(* Logix 5000 project; controller _GigaDiscovery vendor 1 type 14 code 244 rev 35.11; software revision 35.03 *)

TASK _10_milli_sec (periodic, rate 10 ms, priority 5, watchdog 500 ms) : Main10ms
TASK MainTask (continuous, watchdog 500 ms) : Input, Alarms, General, Pylon, Recipe, Output, HMI, Restraints
TASK Pylon_Control (periodic, rate 5 ms, priority 2, watchdog 500 ms) : Pylon_Oscillation
TASK SafetyTask (periodic, rate 40 ms, priority 2, watchdog 20 ms) : S_Input, S_Alarms, S_Cycles, S_Platform_and_Gates, S_Restraints_Release, S_Output

MODULES
   Local : vendor 1 type 14 code 244 (5069 0, rev 35.11)
      Gondola_Motor_7 : vendor 1 type 152 code 121 (Ethernet 192.168.1.63, rev 7.3, Output RPI 20 ms)
           K205_MCC:12:I.4   // Compressor Motor Protection Feedback -F18002C
           K205_MCC:12:I.3   // Compressor Motor Command Feedback -F18101E
           K205_MCC:12:I.2   // Motor 7 Thermal Probe -K16602H
           K205_MCC:12:I.1   // Motor 7 Fan Protection Feedback -F16402C
           K205_MCC:12:I.0   // Zero Set Sensor -B11201A
           K205_MCC:12:I.6   // Platform closed Sector 1 -B22501J
           K205_MCC:12:I.5   // Dryer Motor Protection Feedback -F18202C
           K205_MCC:12:I.7   // Platform closed Sector 2 -B22507J
           K205_MCC:15:I.2   // Magnalock Gate 1 - Status Lock -A25201I
           K205_MCC:15:I.3   // Magnalock Gate 2 - Status Lock -A25207I
           K205_MCC:15:I.4   // Magnalock Gate 3 - Status Lock -A25301I
           K205_MCC:15:I.6   // Feedback Fuse Gondola Motor Power Supply -F16002F -F16003F
           K205_MCC:15:I.7   // Gondola Communication Modem Fault CH1 -T27002C
           K205_MCC:15:I.5   // Magnalock Gate 4 - Status Lock -A25307I
           K205_MCC:15:I.0   // Gate 3 RFID Sensor Closed -B24701J
           K205_MCC:15:I.1   // Gate 4 RFID Sensor Closed -B24801J
           K520_GSB:5:I.0   // Set Number 6
           K520_GSB:5:I.1   // Set Number 7
           K520_GSB:5:I.2   // Set Number 8
           K520_GSB:5:I.3   // Set Number 9
           K520_GSB:5:I.4   // Set Number 10
           K540_GSC:5:I.0   // Set Number 11
           K540_GSC:5:I.1   // Set Number 12
           K540_GSC:5:I.2   // Set Number 13
           K540_GSC:5:I.3   // Set Number 14
           K540_GSC:5:I.4   // Set Number 15
           K600_GSF:5:I.0   // Set Number 26
           K600_GSF:5:I.1   // Set Number 27
           K600_GSF:5:I.2   // Set Number 28
           K600_GSF:5:I.3   // Set Number 29
           K600_GSF:5:I.4   // Set Number 30
           K205_MCC:16:I.0   // Gondola Communication Modem Fault CH2 -T27002C
           K205_MCC:16:I.2   // Fan Feedback NC Pag.94
           K205_MCC:16:I.3   // Fan Feedback NO Pag.94
           K205_MCC:14:I.0   // Platform Opened Sector 3 -B23601J
           K205_MCC:14:I.1   // Platform Opened Sector 4 -B23607J
           K205_MCC:14:I.2   // Platform Opened Sector 5 -B23701J
           K205_MCC:14:I.3   // Platform Opened Sector 6 -B23707J
           K205_MCC:14:I.4   // Platform Opened Sector 7 -B23801J
           K205_MCC:14:I.5   // Platform Opened Sector 8 -B23807J
           K205_MCC:14:I.6   // Gate 1 RFID Sensor Closed -B24501J
           K205_MCC:14:I.7   // Gate 2 RFID Sensor Closed -B24601J
           K205_MCC:11:I.1   // Motor 3 Thermal Probe -K12702H
           K205_MCC:11:I.2   // Motor 4 Thermal Probe -K12704H
           K205_MCC:11:I.6   // Motor 5 Thermal Probe -K14702H
           K205_MCC:11:I.7   // Motor 6 Thermal Probe -K14704H
           K205_MCC:11:I.3   // Motor 5 Overvoltage control - Relay OK -K14302G
           K205_MCC:11:I.4   // Motor 6 Overvoltage control - Relay OK -K14307G
           K205_MCC:11:I.0   // Motor 3-4 Fan Protection Feedback -F12402C -F12406C
           K205_MCC:11:I.5   // Motor 5-6 Fan Protection Feedback -F14402C -F14406C
           K208_MCC:4:O.2   // External Interface Dispatch Command Issued -Q25703H.1
           K208_MCC:4:O.1   // External Interface Automatic Mode -Q25703H
           K208_MCC:4:O.4   // External Interface RCS Fault Status -Q25705H
           K208_MCC:4:O.0   // External Interface Emergency Stop Active -Q25701I
           K208_MCC:4:O.3   // External Interface Fire Alarm -Q25704H
           K208_MCC:4:O.5   // Ride Cycle duration
           K580_GSE:5:I.0   // Set Number 21
           K580_GSE:5:I.1   // Set Number 22
           K580_GSE:5:I.2   // Set Number 23
           K580_GSE:5:I.3   // Set Number 24
           K580_GSE:5:I.4   // Set Number 25
           K205_MCC:17:O.3   // Allow Main Operator OCC2 CONFIRM -S286002F
           K205_MCC:17:O.1   // Fron leg and front light signal -K3204H
           K205_MCC:17:O.7   // UPS MCC
           K205_MCC:17:O.4   // Stop Cycle OCC2 Lamp -S28606F
           K205_MCC:17:O.0   // Rear leg and rear light signal -K3202H
           K205_MCC:17:O.2   // Gondola and pendulum light signal -K3206H
           K205_MCC:17:O.5   // SL RESTRAINTS RELEASE -S28507F
           K205_MCC:17:O   // LIGHT -Q28611I
           K205_MCC:13:I.0   // Platform closed Sector 3 -B22601J
           K205_MCC:13:I.1   // Platform closed Sector 4 -B22607J
           K205_MCC:13:I.2   // Platform closed Sector 5 -B22701J
           K205_MCC:13:I.3   // Platform closed Sector 6 -B22707J
           K205_MCC:13:I.4   // Platform closed Sector 7 -B22801J
           K205_MCC:13:I.5   // Platform closed Sector 8 -B22807J
           K205_MCC:13:I.6   // Platform Opened Sector 1 -B23501J
           K205_MCC:13:I.7   // Platform Opened Sector 2 -B23507J
           K205_MCC:10:I.0   // Motor 1 Overvoltage control - Relay OK -K10302G
           K205_MCC:10:I.1   // Motor 2 Overvoltage control - Relay OK -K10307G
           K205_MCC:10:I.6   // Motor 3 Overvoltage control - Relay OK -K12302G
           K205_MCC:10:I.5   // Pylon Brake Command Feedback -Q10801E
           K205_MCC:10:I.3   // Motor 1 Thermal Probe -K10702H
           K205_MCC:10:I.4   // Motor 2 Thermal Probe -K10704H
           K205_MCC:10:I.7   // Motor 4 Overvoltage control - Relay OK -K12307G
           K205_MCC:10:I.2   // Motor 1-2 Fan Protection Feedback -F10402C -F10406C
           K300_OCC:5:O.0   // .
           K300_OCC:5:O.1   // .
           K300_OCC:5:O.2   // .
           K300_OCC:5:O.3   // .
           K300_OCC:5:O.4   // .
           K300_OCC:5:O.5   // .
           K300_OCC:5:O.6   // .
           K300_OCC:5:O.7   // .
           K620_GSG:5:I.0   // Set Number 31
           K620_GSG:5:I.1   // Set Number 32
           K620_GSG:5:I.2   // Set Number 33
           K620_GSG:5:I.3   // Set Number 34
           K620_GSG:5:I.4   // Set Number 35
           K300_OCC:6:O.3   // +OCC2 -S28502F EMERGENCY
           K300_OCC:6:O.1   // ALARMS BUZZER -P30810F
           K300_OCC:6:O.5   // PLATFORM STOP -S30608F
           K300_OCC:6:O.2   // RESTRAINTS RELEASE Signal Light -S30505F
           K300_OCC:6:O.0   // RESET FAULTS LAMP -S30807F
           K300_OCC:4:I.0   // .
           K300_OCC:4:I.1   // .
           K300_OCC:4:I.2   // .
           K300_OCC:4:I.4   // .
           K500_GSA:5:I.0   // Set Number 1
           K500_GSA:5:I.1   // Set Number 2
           K500_GSA:5:I.2   // Set Number 3
           K500_GSA:5:I.3   // Set Number 4
           K500_GSA:5:I.4   // Set Number 5
           K560_GSD:5:I.0   // Set Number 16
           K560_GSD:5:I.1   // Set Number 17
           K560_GSD:5:I.2   // Set Number 18
           K560_GSD:5:I.3   // Set Number 19
           K560_GSD:5:I.4   // Set Number 20
           K208_MCC:5:O.3   // Load Gate Open Request -Q25904H
           K208_MCC:5:O.2   // Horn -Q25903H.1
           K208_MCC:5:O.1   // Ride Stopping -Q25903H
           K208_MCC:5:O.0   // Ride Stop Active -Q25901
           K640_GSH:5:I.0   // Set Number 36
           K640_GSH:5:I.1   // Set Number 37
           K640_GSH:5:I.2   // Set Number 38
           K640_GSH:5:I.3   // Set Number 39
           K640_GSH:5:I.4   // Set Number 40
          : vendor 1 type 152 code 11008 (DPI 5, rev 1.8)
          : vendor 1 type 152 code 767 (DPI 1, rev 2.7)
      Pylon_Motor_5_6 : vendor 1 type 152 code 121 (Ethernet 192.168.1.62, rev 7.1, Output RPI 20 ms)
          : vendor 1 type 152 code 767 (DPI 1, rev 2.7)
          : vendor 1 type 152 code 11008 (DPI 5, rev 1.4)
      Pylon_Motor_3_4 : vendor 1 type 152 code 121 (Ethernet 192.168.1.61, rev 7.1, Output RPI 20 ms)
          : vendor 1 type 152 code 767 (DPI 1, rev 2.7)
          : vendor 1 type 152 code 11008 (DPI 5, rev 1.4)
      Pylon_Motor_1_2 : vendor 1 type 152 code 121 (Ethernet 192.168.1.60, rev 7.1, Output RPI 20 ms)
           Pylon_Motor_1_2:O.SpdTrqModeSel   // 1 : Speed 2 Torque
          : vendor 1 type 152 code 767 (DPI 1, rev 2.7)
          : vendor 1 type 152 code 11008 (DPI 5, rev 1.4)
      _K20001 : vendor 1 type 109 code 90 (5069 1, rev 3.1, StandardDataDriven RPI 2 ms)
      K300_OCC : 1734-AENTR (Ethernet 192.168.1.10, rev 7.11, Output RPI 20 ms)
           K300_OCC:I.Data[4].1   // Light Selector Switch -S30408F
           K300_OCC:I.Data[4].2   // Reset Status Enable Key -S30801F
           K300_OCC:I.Data[4].0   // Horn Pushbutton -S30407F
           K300_OCC:I.Data[4].4   // OCC Reset Button -S30807F
           K300_OCC:O.Data[5].6   // Platform Close Signal -S30605F
           K300_OCC:O.Data[5].4   // Lapbars open signal -P30509F
           K300_OCC:O.Data[5].3   // Lapbars close signal -P30507F
           K300_OCC:O.Data[5].5   // Platform Open Signal -S30601F
           K300_OCC:O.Data[6].0   // Alarm Lamp -P30810F
           K300_OCC:O.Data[6].1   // Alarm Buzzer -P30810F
           K300_OCC:O.Data[5].0   // Stop Cycle Lamp -S30308F
           K300_OCC:O.Data[5].1   // Start Cycle Lamp -S30403F
           K300_OCC:O.Data[5].2   // Lights On Signal -S30408F
           K300_OCC:O.Data[5].7   // Reset Status Lamp -S30803F
         K30004B : 1734-IB8 (PointIO 4, rev 3.22)
         K30005B : 1734-OB8E (PointIO 5, rev 3.22)
         K30006B : 1734-OB8E (PointIO 6, rev 3.22)
         K30001B : vendor 1 type 35 code 15 (PointIO 1, rev 2.3, Input RPI 35 ms)
              K300_OCC:1:I.Pt02Data   // Operator Enable On/Off
         K30003B : vendor 1 type 35 code 15 (PointIO 3, rev 2.3, Input RPI 35 ms)
         K30002B : vendor 1 type 35 code 15 (PointIO 2, rev 2.3, Input RPI 35 ms)
      K640_GSH : 1734-AENTR (Ethernet 192.168.1.22, rev 5.15, Output RPI 20 ms)
         _05C3 : 1734-IB8 (PointIO 5, rev 3.22)
         _01C3 : vendor 1 type 35 code 15 (PointIO 1, rev 2.3, Input RPI 10 ms, Output RPI 40 ms)
              K640_GSH:1:O.Test02Data   // RFID Supply
         _02C3 : vendor 1 type 35 code 15 (PointIO 2, rev 2.3, Input RPI 10 ms, Output RPI 40 ms)
              K640_GSH:2:O.Test03Data   // RFID Supply
              K640_GSH:2:O.Test00Data   // RFID Supply
              K640_GSH:2:O.Test02Data   // RFID Supply
              K640_GSH:2:O.Test01Data   // RFID Supply
         _04C3 : vendor 1 type 35 code 16 (PointIO 4, rev 2.3, Output RPI 40 ms, Input RPI 35 ms)
              K640_GSH:4:O.Pt05Data   // Right Rack Unlick Valve -B46005I
              K640_GSH:4:O.Pt07Data   // Left Rack Unlock Valve -B47002I
              K640_GSH:4:O.Pt01Data   // Right Rack Unlock Valve -B64505I
              K640_GSH:4:O.Pt02Data   // LAPBARS OPENING VALVE -B64508I
              K640_GSH:4:O.Pt00Data   // Left Rack Unlock Valve -B64502I
              K640_GSH:4:O.Pt04Data   // Left Rack Unlick Valve -B46002I
              K640_GSH:4:O.Pt03Data   // Open Valve -B45008I
              K640_GSH:4:O.Pt06Data   // Open Valve -B46008I
         _03C3 : vendor 1 type 35 code 15 (PointIO 3, rev 2.1, Input RPI 10 ms, Output RPI 40 ms)
              K640_GSH:3:O.Test03Data   // RFID Supply
              K640_GSH:3:O.Test00Data   // RFID Supply
              K640_GSH:3:O.Test02Data   // RFID Supply
              K640_GSH:3:O.Test01Data   // RFID Supply
      K500_GSA : 1734-AENTR (Ethernet 192.168.1.14, rev 5.15, Output RPI 20 ms)
         K39505C : 1734-IB8 (PointIO 5, rev 3.22)
         K39502C : vendor 1 type 35 code 15 (PointIO 2, rev 2.3, Output RPI 40 ms, Input RPI 10 ms)
              K500_GSA:2:O.Test03Data   // RFID Supply
              K500_GSA:2:O.Test00Data   // RFID Supply
              K500_GSA:2:O.Test02Data   // RFID Supply
              K500_GSA:2:O.Test01Data   // RFID Supply
         K50001C : vendor 1 type 35 code 15 (PointIO 3, rev 2.1, Output RPI 40 ms, Input RPI 10 ms)
              K500_GSA:3:O.Test03Data   // RFID Supply
              K500_GSA:3:O.Test00Data   // RFID Supply
              K500_GSA:3:O.Test02Data   // RFID Supply
              K500_GSA:3:O.Test01Data   // RFID Supply
         K39501C : vendor 1 type 35 code 15 (PointIO 1, rev 2.3, Input RPI 10 ms, Output RPI 40 ms)
              K500_GSA:1:O.Test02Data   // RFID Supply
         K39503C : vendor 1 type 35 code 16 (PointIO 4, rev 2.3, Output RPI 40 ms, Input RPI 35 ms)
              K500_GSA:4:O.Pt00Data   // Right Rack Unlock Valve -B50502I
              K500_GSA:4:O.Pt07Data   // Left Rack Unlock Valve -B47002I
              K500_GSA:4:O.Pt05Data   // Right Rack Unlick Valve -B46005I
              K500_GSA:4:O.Pt01Data   // Left Rack Unlock Valve -B50505I
              K500_GSA:4:O.Pt04Data   // Left Rack Unlick Valve -B46002I
              K500_GSA:4:O.Pt02Data   // LAPBARS OPENING VALVE -B50508I
              K500_GSA:4:O.Pt03Data   // Open Valve -B45008I
              K500_GSA:4:O.Pt06Data   // Open Valve -B46008I
      K560_GSD : 1734-AENTR (Ethernet 192.168.1.17, rev 5.15, Output RPI 20 ms)
         _05C11 : 1734-IB8 (PointIO 5, rev 3.22)
         _04C11 : vendor 1 type 35 code 16 (PointIO 4, rev 2.3, Input RPI 35 ms, Output RPI 40 ms)
              K560_GSD:4:O.Pt02Data   // LAPBARS OPENING VALVE -B56208I
              K560_GSD:4:O.Pt07Data   // Left Rack Unlock Valve -B47002I
              K560_GSD:4:O.Pt00Data   // Left Rack Unlock Valve -B56202I
              K560_GSD:4:O.Pt05Data   // Right Rack Unlick Valve -B46005I
              K560_GSD:4:O.Pt01Data   // Right Rack Unlock Valve -B56205I
              K560_GSD:4:O.Pt04Data   // Left Rack Unlick Valve -B46002I
              K560_GSD:4:O.Pt03Data   // Open Valve -B45008I
              K560_GSD:4:O.Pt06Data   // Open Valve -B46008I
         _03C11 : vendor 1 type 35 code 15 (PointIO 3, rev 2.1, Output RPI 40 ms, Input RPI 10 ms)
              K560_GSD:3:O.Test03Data   // RFID Supply
              K560_GSD:3:O.Test00Data   // RFID Supply
              K560_GSD:3:O.Test02Data   // RFID Supply
              K560_GSD:3:O.Test01Data   // RFID Supply
         _01C11 : vendor 1 type 35 code 15 (PointIO 1, rev 2.3, Input RPI 10 ms, Output RPI 40 ms)
              K560_GSD:1:O.Test02Data   // RFID Supply
         _02C11 : vendor 1 type 35 code 15 (PointIO 2, rev 2.3, Input RPI 10 ms, Output RPI 40 ms)
              K560_GSD:2:O.Test03Data   // RFID Supply
              K560_GSD:2:O.Test00Data   // RFID Supply
              K560_GSD:2:O.Test02Data   // RFID Supply
              K560_GSD:2:O.Test01Data   // RFID Supply
      K390_GMB_RCC1 : 1734-AENTR (Ethernet 192.168.1.13, rev 5.15, Output RPI 20 ms)
         K39007C : 1734-IB8 (PointIO 4, rev 3.22)
         K39004C : vendor 1 type 35 code 16 (PointIO 3, rev 2.3, Output RPI 40 ms, Input RPI 35 ms)
              K390_GMB_RCC1:3:O.Pt03Data   // Open Valve -B41008I
              K390_GMB_RCC1:3:O.Pt07Data   // Left Rack Unlock Valve -B43002I
              K390_GMB_RCC1:3:O.Pt04Data   // Left Rack Unlock Valve -B42002I
              K390_GMB_RCC1:3:O.Pt05Data   // Right Rack Unlock Valve -B42005I
              K390_GMB_RCC1:3:O.Pt00Data   // Main Valve -B40501I
              K390_GMB_RCC1:3:O.Pt06Data   // Open Valve -B42008I
              K390_GMB_RCC1:3:O.Pt02Data   // Horn -P40702I
         K39001C : vendor 1 type 35 code 15 (PointIO 1, rev 2.3, Input RPI 35 ms)
              K390_GMB_RCC1:1:I.Pt05Data   // Main Valve Close Limit Switch -B40508I
              K390_GMB_RCC1:1:I.Pt04Data   // Main Valve Open Limit Switch -B40504I
              K390_GMB_RCC1:1:I.Pt02Data   // +GMB_RCC1 Temperature OK -S40103E
              K390_GMB_RCC1:1:I.Pt00Data   // Home Sensor Speed Check -B40002I
              K390_GMB_RCC1:1:I.Pt01Data   // Home Sensor Speed Check -B40007I
         K39002C : vendor 1 type 35 code 15 (PointIO 2, rev 2.3, Input RPI 35 ms)
              K390_GMB_RCC1:2:I.Pt05Data   // +RCC_GSF Temperature OK -S60110G
              K390_GMB_RCC1:2:I.Pt01Data   // +RCC_GSB Temperature OK -S52110G
              K390_GMB_RCC1:2:I.Pt07Data   // +RCC_GSH Temperature OK -S64110G
              K390_GMB_RCC1:2:I.Pt00Data   // +RCC_GSA Temperature OK -S50110G
              K390_GMB_RCC1:2:I.Pt04Data   // +RCC_GSE Temperature OK -S58110G
              K390_GMB_RCC1:2:I.Pt06Data   // +RCC_GSG Temperature OK -S62110G
              K390_GMB_RCC1:2:I.Pt03Data   // +RCC_GSD Temperature OK -S56110G
              K390_GMB_RCC1:2:I.Pt02Data   // +RCC_GSC Temperature OK -S54110G
      K540_GSC : 1734-AENTR (Ethernet 192.168.1.16, rev 5.15, Output RPI 20 ms)
         _05C1 : 1734-IB8 (PointIO 5, rev 3.22)
         _02C1 : vendor 1 type 35 code 15 (PointIO 2, rev 2.3, Input RPI 10 ms, Output RPI 40 ms)
              K540_GSC:2:O.Test03Data   // RFID Supply
              K540_GSC:2:O.Test00Data   // RFID Supply
              K540_GSC:2:O.Test02Data   // RFID Supply
              K540_GSC:2:O.Test01Data   // RFID Supply
         _04C1 : vendor 1 type 35 code 16 (PointIO 4, rev 2.3, Input RPI 35 ms, Output RPI 40 ms)
              K540_GSC:4:O.Pt02Data   // LAPBARS OPENING VALVE -B54508I
              K540_GSC:4:O.Pt07Data   // Left Rack Unlock Valve -B47002I
              K540_GSC:4:O.Pt01Data   // Left Rack Unlock Valve -B54502I
              K540_GSC:4:O.Pt03Data   // Open Valve -B45008I
              K540_GSC:4:O.Pt06Data   // Open Valve -B46008I
              K540_GSC:4:O.Pt04Data   // Left Rack Unlick Valve -B46002I
              K540_GSC:4:O.Pt00Data   // Right Rack Unlock Valve -B54505I
              K540_GSC:4:O.Pt05Data   // Right Rack Unlick Valve -B46005I
         _03C1 : vendor 1 type 35 code 15 (PointIO 3, rev 2.1, Input RPI 10 ms, Output RPI 40 ms)
              K540_GSC:3:O.Test00Data   // RFID Supply
              K540_GSC:3:O.Test01Data   // RFID Supply
         _01C1 : vendor 1 type 35 code 15 (PointIO 1, rev 2.3, Input RPI 10 ms, Output RPI 40 ms)
              K540_GSC:1:O.Test02Data   // RFID Supply
      K620_GSG : 1734-AENTR (Ethernet 192.168.1.20, rev 5.15, Output RPI 20 ms)
         _05C2 : 1734-IB8 (PointIO 5, rev 3.22)
         _02C2 : vendor 1 type 35 code 15 (PointIO 2, rev 2.3, Input RPI 10 ms, Output RPI 40 ms)
              K620_GSG:2:O.Test03Data   // RFID Supply
              K620_GSG:2:O.Test00Data   // RFID Supply
              K620_GSG:2:O.Test02Data   // RFID Supply
              K620_GSG:2:O.Test01Data   // RFID Supply
         _01C2 : vendor 1 type 35 code 15 (PointIO 1, rev 2.3, Input RPI 10 ms, Output RPI 40 ms)
              K620_GSG:1:O.Test02Data   // RFID Supply
         _04C2 : vendor 1 type 35 code 16 (PointIO 4, rev 2.3, Input RPI 35 ms, Output RPI 40 ms)
              K620_GSG:4:O.Pt05Data   // Right Rack Unlick Valve -B46005I
              K620_GSG:4:O.Pt07Data   // Left Rack Unlock Valve -B47002I
              K620_GSG:4:O.Pt01Data   // Right Rack Unlock Valve -B62505I
              K620_GSG:4:O.Pt00Data   // Left Rack Unlock Valve -B62502I
              K620_GSG:4:O.Pt04Data   // Left Rack Unlick Valve -B46002I
              K620_GSG:4:O.Pt02Data   // LAPBARS OPENING VALVE -B62508I
              K620_GSG:4:O.Pt03Data   // Open Valve -B45008I
              K620_GSG:4:O.Pt06Data   // Open Valve -B46008I
         _03C2 : vendor 1 type 35 code 15 (PointIO 3, rev 2.1, Input RPI 10 ms, Output RPI 40 ms)
              K620_GSG:3:O.Test03Data   // RFID Supply
              K620_GSG:3:O.Test00Data   // RFID Supply
              K620_GSG:3:O.Test02Data   // RFID Supply
              K620_GSG:3:O.Test01Data   // RFID Supply
      K580_GSE : 1734-AENTR (Ethernet 192.168.1.18, rev 5.15, Output RPI 20 ms)
         _05C111 : 1734-IB8 (PointIO 5, rev 3.22)
         _04C111 : vendor 1 type 35 code 16 (PointIO 4, rev 2.3, Output RPI 40 ms, Input RPI 35 ms)
              K580_GSE:4:O.Pt02Data   // LAPBARS OPENING VALVE -B58508I
              K580_GSE:4:O.Pt07Data   // Left Rack Unlock Valve -B47002I
              K580_GSE:4:O.Pt00Data   // Left Rack Unlock Valve -B58502I
              K580_GSE:4:O.Pt04Data   // Left Rack Unlick Valve -B46002I
              K580_GSE:4:O.Pt05Data   // Right Rack Unlick Valve -B46005I
              K580_GSE:4:O.Pt01Data   // Right Rack Unlock Valve -B58505I
              K580_GSE:4:O.Pt03Data   // Open Valve -B45008I
              K580_GSE:4:O.Pt06Data   // Open Valve -B46008I
         _03C111 : vendor 1 type 35 code 15 (PointIO 3, rev 2.1, Output RPI 40 ms, Input RPI 10 ms)
              K580_GSE:3:O.Test03Data   // RFID Supply
              K580_GSE:3:O.Test00Data   // RFID Supply
              K580_GSE:3:O.Test02Data   // RFID Supply
              K580_GSE:3:O.Test01Data   // RFID Supply
         _02C111 : vendor 1 type 35 code 15 (PointIO 2, rev 2.3, Input RPI 10 ms, Output RPI 40 ms)
              K580_GSE:2:O.Test03Data   // RFID Supply
              K580_GSE:2:O.Test00Data   // RFID Supply
              K580_GSE:2:O.Test02Data   // RFID Supply
              K580_GSE:2:O.Test01Data   // RFID Supply
         _01C111 : vendor 1 type 35 code 15 (PointIO 1, rev 2.3, Input RPI 10 ms, Output RPI 40 ms)
              K580_GSE:1:O.Test02Data   // RFID Supply
      K520_GSB : 1734-AENTR (Ethernet 192.168.1.15, rev 5.15, Output RPI 20 ms)
         _05C : 1734-IB8 (PointIO 5, rev 3.22)
         _01C : vendor 1 type 35 code 15 (PointIO 1, rev 2.3, Output RPI 40 ms, Input RPI 10 ms)
              K520_GSB:1:O.Test02Data   // RFID Supply
         _04C : vendor 1 type 35 code 16 (PointIO 4, rev 2.3, Output RPI 40 ms, Input RPI 35 ms)
              K520_GSB:4:O.Pt02Data   // LAPBARS OPENING VALVE -B52508I
              K520_GSB:4:O.Pt07Data   // Left Rack Unlock Valve -B47002I
              K520_GSB:4:O.Pt01Data   // Left Rack Unlock Valve -B52502I
              K520_GSB:4:O.Pt04Data   // Left Rack Unlick Valve -B46002I
              K520_GSB:4:O.Pt00Data   // Right Rack Unlock Valve -B52505I
              K520_GSB:4:O.Pt03Data   // Open Valve -B45008I
              K520_GSB:4:O.Pt06Data   // Open Valve -B46008I
              K520_GSB:4:O.Pt05Data   // Right Rack Unlick Valve -B46005I
         _02C : vendor 1 type 35 code 15 (PointIO 2, rev 2.3, Output RPI 40 ms, Input RPI 10 ms)
              K520_GSB:2:O.Test03Data   // RFID Supply
              K520_GSB:2:O.Test00Data   // RFID Supply
              K520_GSB:2:O.Test02Data   // RFID Supply
              K520_GSB:2:O.Test01Data   // RFID Supply
         _03C : vendor 1 type 35 code 15 (PointIO 3, rev 2.1, Input RPI 10 ms, Output RPI 40 ms)
              K520_GSB:3:O.Test03Data   // RFID Supply
              K520_GSB:3:O.Test00Data   // RFID Supply
              K520_GSB:3:O.Test02Data   // RFID Supply
              K520_GSB:3:O.Test01Data   // RFID Supply
      K600_GSF : 1734-AENTR (Ethernet 192.168.1.19, rev 7.11, Output RPI 20 ms)
         _05C1111 : 1734-IB8 (PointIO 5, rev 3.31)
         _03C1111 : vendor 1 type 35 code 15 (PointIO 3, rev 2.1, Input RPI 10 ms, Output RPI 40 ms)
              K600_GSF:3:O.Test03Data   // RFID Supply
              K600_GSF:3:O.Test00Data   // RFID Supply
              K600_GSF:3:O.Test02Data   // RFID Supply
              K600_GSF:3:O.Test01Data   // RFID Supply
         _02C1111 : vendor 1 type 35 code 15 (PointIO 2, rev 2.3, Input RPI 10 ms, Output RPI 40 ms)
              K600_GSF:2:O.Test03Data   // RFID Supply
              K600_GSF:2:O.Test00Data   // RFID Supply
              K600_GSF:2:O.Test02Data   // RFID Supply
              K600_GSF:2:O.Test01Data   // RFID Supply
         _04C1111 : vendor 1 type 35 code 16 (PointIO 4, rev 2.3, Input RPI 35 ms, Output RPI 40 ms)
              K600_GSF:4:O.Pt07Data   // Left Rack Unlock Valve -B47002I
              K600_GSF:4:O.Pt01Data   // Left Rack Unlock Valve -B60505I
              K600_GSF:4:O.Pt04Data   // Left Rack Unlick Valve -B46002I
              K600_GSF:4:O.Pt00Data   // Right Rack Unlock Valve -B60502I
              K600_GSF:4:O.Pt05Data   // Right Rack Unlick Valve -B46005I
              K600_GSF:4:O.Pt02Data   // LAPBARS OPENING VALVE -B60508I
              K600_GSF:4:O.Pt03Data   // Open Valve -B45008I
              K600_GSF:4:O.Pt06Data   // Open Valve -B46008I
         _01C1111 : vendor 1 type 35 code 15 (PointIO 1, rev 2.3, Output RPI 40 ms, Input RPI 10 ms)
              K600_GSF:1:O.Test02Data   // RFID Supply
      K205_MCC : 1734-AENTR (Ethernet 192.168.1.11, rev 7.11, Output RPI 20 ms)
         K20515C : 1734-IB8 (PointIO 15, rev 3.22)
         K20512C : 1734-IB8 (PointIO 12, rev 3.22)
         K20516C : 1734-IB8 (PointIO 16, rev 3.22)
         K20511C : 1734-IB8 (PointIO 11, rev 3.22)
         K20514C : 1734-IB8 (PointIO 14, rev 3.22)
         K20510C : 1734-IB8 (PointIO 10, rev 3.22)
         K20513C : 1734-IB8 (PointIO 13, rev 3.22)
         K20517C : 1734-OB8E (PointIO 17, rev 3.22)
         K20502C : vendor 1 type 35 code 15 (PointIO 2, rev 2.3, Input RPI 10 ms)
              K205_MCC:2:I.Pt02Data   // Platform Close Main Valve Limit Switch -B21909I
              K205_MCC:2:I.Pt00Data   // Platform Line Minimum Pressure Switch -S21511B
              K205_MCC:2:I.Pt01Data   // Platform Open Main Valve Limit Switch -B21905I
         K20506C : vendor 1 type 35 code 15 (PointIO 6, rev 2.3, Input RPI 35 ms)
         K20501C : vendor 1 type 35 code 15 (PointIO 1, rev 2.3, Input RPI 35 ms)
              K205_MCC:1:I.Pt03Data   // Gondola Motor - Start Feedback -Q16105E -Q16107E -Q16202G
              K205_MCC:1:I.Pt04Data   // Line Pressure Switch - Working Pressure -S21502B
              K205_MCC:1:I.Pt05Data   // Line Pressure Switch - Minimum Pressure -S21504B
              K205_MCC:1:I.Pt06Data   // Platform Maximum Opening Pressure -S21507B
              K205_MCC:1:I.Pt07Data   // Platform Maximum Closing Pressure -S21510B
         K20507C : vendor 1 type 35 code 16 (PointIO 7, rev 2.3, Input RPI 35 ms, Output RPI 40 ms)
              K205_MCC:7:O.Pt05Data   // Brake Emergency Valve Motor 5 -Y22102I
              K205_MCC:7:O.Pt06Data   // Brake Emergency Valve Motor 6 -Y22108I
              K205_MCC:7:O.Pt03Data   // Pylon Drive 1-2 Start Contactor -Q9002H
              K205_MCC:7:O.Pt00Data   // Pylon Drive Field Contactor -Q10101E
              K205_MCC:7:O.Pt04Data   // Pylon Drive 1-2 Start Contactor -Q9004H
              K205_MCC:7:O.Pt07Data   // Gondola Motor Command -Q16101E
              K205_MCC:7:O.Pt02Data   // Pylon Brake Command -Q10801E
              K205_MCC:7:O.Pt01Data   // Pylon Drive Field Contactor -Q10103E
         K20518C : vendor 1 type 35 code 16 (PointIO 18, rev 2.3, Input RPI 35 ms, Output RPI 40 ms)
              K205_MCC:18:O.Pt01Data   // Gondola Drive Enable Ch1 Contactor -Q16105E
              K205_MCC:18:O.Pt05Data   // Pylon Drive 3 -4 Start Contactor -Q9007E
              K205_MCC:18:O.Pt07Data   // Pylon Drive 5 - 6 Start Contactor -Q9011E
              K205_MCC:18:O.Pt02Data   // Gondola Drive Enable Ch2 Contactor -Q16107E
              K205_MCC:18:O.Pt00Data   // Pilot Valves Enable for Opening/Closing Platform - Y22002A
              K205_MCC:18:O.Pt04Data   // Pylon Drive 3 - 4 Start Contactor -Q9005E
              K205_MCC:18:O.Pt06Data   // Pylon Drive 5 - 6 Start Contactor -Q9009E
              K205_MCC:18:O.Pt03Data   // Pylon Motors Fan -Q9302F
         K20508C : vendor 1 type 35 code 16 (PointIO 8, rev 2.3, Input RPI 35 ms, Output RPI 40 ms)
              K205_MCC:8:O.Pt00Data   // Gondola Motor Command -Q16103E
              K205_MCC:8:O.Pt06Data   // Valvola principale piattaforma B21902I
              K205_MCC:8:O.Pt03Data   // Platform Opening Valve -Y21706I
              K205_MCC:8:O.Pt05Data   // Platform Opening Valve -Y21806I
              K205_MCC:8:O.Pt04Data   // Platform Closing Valve -Y21802I
              K205_MCC:8:O.Pt02Data   // Platform Closing Valve -Y21702I
              K205_MCC:8:O.Pt07Data   // Gate Lock Enable -Q25102E
         K20505C : vendor 1 type 35 code 15 (PointIO 5, rev 2.3, Input RPI 10 ms)
         K20504C : vendor 1 type 35 code 15 (PointIO 4, rev 2.3, Input RPI 35 ms)
              K205_MCC:4:I.Pt02Data   // Unlock Platform Line Pressure Switch -S22006B
              K205_MCC:4:I.Pt05Data   // MCC temeprature OK -S75003C
         K20503C : vendor 1 type 35 code 15 (PointIO 3, rev 2.3, Output RPI 40 ms, Input RPI 35 ms)
              K205_MCC:3:O.Test03Data   // Reset RFID Platform Closed Sensors Page 225
              K205_MCC:3:O.Test01Data   // Reset Gate RFID Sensor -B24501J ... -B24802J
              K205_MCC:3:O.Test02Data   // Reset RFID Platform Opened Sensors Page 2
         K20509C : vendor 1 type 42 code 1 (PointIO 9, rev 1.3, Output RPI 40 ms, Input RPI 35 ms)
      K208_MCC : 1734-AENTR (Ethernet 192.168.1.12, rev 6.13, Output RPI 20 ms)
         K20804C : 1734-OB8 (PointIO 4, rev 3.1)
         K20805C : 1734-OB8 (PointIO 5, rev 3.1)
         K20803C : vendor 1 type 35 code 15 (PointIO 3, rev 2.3, Input RPI 10 ms, Output RPI 40 ms)
              K208_MCC:3:I.Pt04Data   // Line Pressure Switch - Working Pressure -S21502B
              K208_MCC:3:I.Pt03Data   // Gondola Motor - Start Feedback -Q16105E -Q16107E -Q16202G
              K208_MCC:3:I.Pt05Data   // Line Pressure Switch - Minimum Pressure -S21504B
              K208_MCC:3:I.Pt06Data   // Platform Maximum Opening Pressure -S21507B
              K208_MCC:3:I.Pt07Data   // Platform Maximum Closing Pressure -S21510B
         K20802C : vendor 1 type 35 code 16 (PointIO 2, rev 2.3, Input RPI 35 ms, Output RPI 40 ms)
              K208_MCC:2:O.Pt05Data   // Brake Emergency Valve Motor 5 -Y22102I
              K208_MCC:2:O.Pt02Data   // Pylon Brake Command -Q10801E
              K208_MCC:2:O.Pt07Data   // Gondola Motor Command -Q16101E
              K208_MCC:2:O.Pt01Data   // Pylon Drive Field Contactor -Q10103E
              K208_MCC:2:O.Pt06Data   // Brake Emergency Valve Motor 6 -Y22108I
              K208_MCC:2:O.Pt03Data   // Pylon Drive 1-2 Start Contactor -Q9002H
              K208_MCC:2:O.Pt04Data   // Pylon Drive 1-2 Start Contactor -Q9004H
         K20801C : vendor 1 type 35 code 15 (PointIO 1, rev 2.3, Input RPI 35 ms)
              K208_MCC:1:I.Pt04Data   // Line Pressure Switch - Working Pressure -S21502B
              K208_MCC:1:I.Pt05Data   // Line Pressure Switch - Minimum Pressure -S21504B
              K208_MCC:1:I.Pt06Data   // Platform Maximum Opening Pressure -S21507B
              K208_MCC:1:I.Pt07Data   // Platform Maximum Closing Pressure -S21510B
END_MODULES

TYPE AssetSettings :
STRUCT
   AssetID : DINT;
   AlarmsOffset : DINT;
END_STRUCT
END_TYPE

TYPE Auto_Cycle :
STRUCT
   Pylon_Angle : DINT;
   Cycle_Time_min : DINT;
   Cycle_Time_sec : DINT;
   Gondola_Speed : DINT[11];
   Gondola_Time : DINT[11];
END_STRUCT
END_TYPE

TYPE Axe :
STRUCT
   Speed : REAL;
   Speed_ABS : REAL;
   Position_0_360 : REAL;
   Position_Sign_180 : REAL;
   Position_Abs_180 : REAL;
END_STRUCT
END_TYPE

TYPE Data_time :
STRUCT
   Year : DINT;
   Month : DINT;
   Day : DINT;
   Hour : DINT;
   Minute : DINT;
   Second : DINT;
   Milli_sec : DINT;
END_STRUCT
END_TYPE

TYPE EventsGroup :
STRUCT
   ActualState : DINT;
   PrevState : DINT;
   ChangedState : DINT;
   RiseEdge : DINT;
   FallEdge : DINT;
   EventID : DINT[32];
   RiseValue : DINT[32];
   FallValue : DINT[32];
END_STRUCT
END_TYPE

TYPE Lap_Bars_Sfty :
STRUCT
   Enable_Unlock_Right_Valve : BOOL;
   Enable_Unlock_Left_Valve : BOOL;
   Lift_Valve : BOOL;
   O_Unlock_Right_Valve : Valve_2_pos_monostable;
   O_Unlock_Left_Valve : Valve_2_pos_monostable;
   I_Down_Position : UDT_DCM;
   I_Sector_Enable : UDT_DCM;
END_STRUCT
END_TYPE

TYPE Lap_Bars_Std :
STRUCT
   Position_Down : BOOL;
   Opened_in_Start_memory : BOOL;
END_STRUCT
END_TYPE

TYPE LapBar_Racks :
STRUCT
   Input_Left : AOI_DCM;
   Input_Right : AOI_DCM;
   ON_Delay_Left : TIMER;
   ON_Delay_Right : TIMER;
   Memory_Left : BOOL;   // Memory Locked
   Memory_Right : BOOL;   // Memory Locked
   Os_Left : BOOL;
   Os_Right : BOOL;
   Memory_Left_Unlocked : BOOL;   // Memory UNLocked
   Memory_Right_Unlocked : BOOL;   // Memory UNLocked
END_STRUCT
END_TYPE

TYPE LapBars_Monitor :
STRUCT
   Sensor_Open_Memory : BOOL;
   Status : BOOL;
END_STRUCT
END_TYPE

TYPE LapBars_Sector :
STRUCT
   Sensors_ChA : BOOL;
   Sensors_ChB : BOOL;
   LapBar_Open_Close : BOOL;
   Input_Status : BOOL;
   Sensor_ChA_Open_Memory : BOOL;
   Sensor_ChB_Open_Memory : BOOL;
   I_LB_PressureSwitch_Valve_Right_Open : BOOL;
   I_LB_PressureSwitch_Valve_Left_Open : BOOL;
   O_LapBars_Valve_Lift : BOOL;
   O_Enable_Unlock_Right_Valve : BOOL;
   O_Enable_Unlock_Left_Valve : BOOL;
   All_Rack_Memory_Signal_ON : BOOL;
   RESTRAINTS_Rack_Sector_ON : BOOL;
   I_Close_Position : DCI_MONITOR;
   I_Sector_Disable_Switch : UDT_DCM;   // 0 = Enabled 1 = Disabled
   O_Unlock_Valve_Left : Valve_2_pos_monostable;
   O_Unlock_Valve_Right : Valve_2_pos_monostable;
END_STRUCT
END_TYPE

TYPE MasterRTUQueue :
STRUCT
   Size : DINT;   // size of array, loaded at startup
   PTR : DINT;   // actual pointer
   Buffer : SERVER_Interface_RTUData[200];
END_STRUCT
END_TYPE

TYPE Permissive :
STRUCT
   All_Permissive_Ok : BOOL;
   BitsConditions : DINT;
   Automatic_I_Stop_Delay : TIMER;
END_STRUCT
END_TYPE

TYPE Permissive_Description :
STRUCT
   OS_Fail : BOOL;
   FailBitsConditions : DINT;
   Visible_Bits : DINT;
   Header_Description_en : STRING;
   Header_Description_others : STRING;
   Bit_Description_en : STRING[32];
   Bit_Description_others : STRING[32];
END_STRUCT
END_TYPE

TYPE PlcClockManaged :
STRUCT
   SetDateTime : BOOL;
   DisableUpdate : BOOL;
   DateTimeValid : BOOL;
   ActualTimestamp_A : DINT;
   ActualTimestamp_B : DINT;
   ActualDateTime : DINT[7];
   DateTimeToSet : DINT[7];
END_STRUCT
END_TYPE

TYPE Proof_Test :
STRUCT
   Left : BOOL;
   Right : BOOL;
   Request : BOOL;
   Reset : BOOL;
   Validation_Delay_time : TIMER;
END_STRUCT
END_TYPE

TYPE Run_Count_Hist_JM :
STRUCT
   date : DINT[3];
   runs : DINT[30];
   time_avg : DINT[30];
END_STRUCT
END_TYPE

TYPE S_Curve_Calc :
STRUCT
   Jerk_Time : REAL;
   Accel_Time : REAL;
   Jerk_Rate : REAL;
   Accel_Rate : REAL;
END_STRUCT
END_TYPE

TYPE Scale_2_P :
STRUCT
   Input : REAL[2];
   Output : REAL[2];
END_STRUCT
END_TYPE

TYPE Sequencer :
STRUCT
   Index : DINT;
   OS : DINT[2];
   Step_Timer : TIMER[32];
   Time_Limit : TIMER[32];
   Alarms_TimeLimit : DINT;
   Started : BOOL;
   Started_OFF_Delay : BOOL;
   Step_00 : BOOL;
   Step_01 : BOOL;
   Step_02 : BOOL;
   Step_03 : BOOL;
   Step_04 : BOOL;
   Step_05 : BOOL;
   Step_06 : BOOL;
   Step_07 : BOOL;
   Step_08 : BOOL;
   Step_09 : BOOL;
   Step_10 : BOOL;
   Step_11 : BOOL;
   Step_12 : BOOL;
   Step_13 : BOOL;
   Step_14 : BOOL;
   Step_15 : BOOL;
   Step_16 : BOOL;
   Step_17 : BOOL;
   Step_18 : BOOL;
   Step_19 : BOOL;
   Step_20 : BOOL;
   Step_21 : BOOL;
   Step_22 : BOOL;
   Step_23 : BOOL;
   Step_24 : BOOL;
   Step_25 : BOOL;
   Step_26 : BOOL;
   Step_27 : BOOL;
   Step_28 : BOOL;
   Step_29 : BOOL;
   Step_30 : BOOL;
   Step_31 : BOOL;
END_STRUCT
END_TYPE

TYPE SERVER_Interface_Ctrl :
STRUCT
   WriteTimeout : TIMER;
   WriteRequest : BOOL;
   HeartBeat : BOOL;
   ReadCompleted : BOOL;
END_STRUCT
END_TYPE

TYPE SERVER_Interface_RTUData :
STRUCT
   LogixID : DINT;
   EventID : DINT;
   DataValue : DINT;
   TimeStamp : Data_time;
END_STRUCT
END_TYPE

TYPE Status_Safety :
STRUCT
   SafetyLockedState : DINT;
   SafetySignatureExists : DINT;
   SafetySignature : STRING;
   Date : STRING;
END_STRUCT
END_TYPE

TYPE Std_to_Sfty :
STRUCT
   Seat_Auxiliary_Ch_Memory : BOOL;
   Gondola_Decc_timer_Start : BOOL;
   I_Fan_Feedback_NC : BOOL;
   I_Fan_Feedback_NO : BOOL;
   Alarms_Reset : BOOL;
   Ride_Stopping : BOOL;
   Stop_Request : BOOL;
   RFID_Reset : BOOL;
   No_Std_Emergencies_CL0 : BOOL;
   No_Std_Emergencies_CL1 : BOOL;
   Ready_to_Stop : BOOL;
   Pylon_min_speed : BOOL;
   Gondola_min_Speed : BOOL;
   Pylon_Stop_at_Home : BOOL;
   Ack_LapBars_ProofTest : BOOL;
   Fbk_MainCotnactor_M1_M3 : BOOL;
   Fbk_MainContactor_M2_M4 : BOOL;
   Fbk_MainContactor_M5 : BOOL;
   Fbk_Compressor_Contactor : BOOL;   // Compressor Motor Command Feedback -F18101E
   Fbk_PylonBrake_Contactor : BOOL;   // Pylon Brake Command Feedback -Q10801E
   I_Magnalock_1_Closed : BOOL;
   I_Magnalock_2_Closed : BOOL;
   I_Magnalock_3_Closed : BOOL;
   I_Magnalock_4_Closed : BOOL;
   I_OCC1_Alarms_Reset_Pb : BOOL;
   I_OCC2_Alarms_Reset_Pb : BOOL;
   HMI_Pb_ProofTest_RESET : BOOL;
   HMI_Bypass_Proof_Test : BOOL;
   Reset_Status : BOOL;
   Horn : BOOL;   // -P40702I
   I_Gondola_Field_Contactor_Fdbk : BOOL;   // Gondola Drive Field Contactors Feedback -Q16101E -Q16103E -Q16202G -Q16202G
   I_Gondola_Fuse_Power_Supply : BOOL;   // Feedback Fuse Gondola Motor Power Supply -F16002F -F16003F
   Pneumatic_Brake_Cmd : BOOL;
   Motors_Temperature_Ok : BOOL;
   Zero_Set_Sensor : BOOL;   // Zero Set Sensor -B11201A
   ACKNOWLEDGE : BOOL;   // ACKNOWLEDGE4 -S30807F
   HMI_Platform_Open : BOOL;
   HMI_Platform_Close : BOOL;
   Low_speed_thold_emergency_brake : BOOL;
   UPS_RCC : UPS;   // -T37603B
   UPS_MCC : UPS;   // -T6603B
   Pylon_Motor_1_3 : Std_to_Sfty_Drive;
   Pylon_Motor_2_4 : Std_to_Sfty_Drive;
   Pylon_Motor_5_6 : Std_to_Sfty_Drive;
   Gondola_Motor_7 : Std_to_Sfty_Drive;
   Gondola_Motor_7ISpdFeedback : DINT;
   Pylon_angle : DINT;
   Main_valve_Time : DINT;
   HMI_Page : DINT;
   HMI_Disable_Opening_Bars : DINT;
   Last_Angle_Reached : REAL;
   Date_Time : Data_time;
   RESTRAINTS_Open_Postion_Aux_Seat : BOOL[64];
END_STRUCT
END_TYPE

TYPE Std_to_Sfty_Drive :
STRUCT
   StopAssert : BOOL;
   Status_Ready : BOOL;
   Status_Active : BOOL;
END_STRUCT
END_TYPE

TYPE UDT_CROUT :
STRUCT
   CROUT : CONFIGURABLE_ROUT;
   Timer : TIMER;
   Actuate : BOOL;
   Out_Status : BOOL;
   In_Status : BOOL;
END_STRUCT
END_TYPE

TYPE UDT_DCI_STOP_TEST :
STRUCT
   Push_Botton : DCI_STOP_TEST;
   Status : BOOL;
   Test_Request : BOOL;
END_STRUCT
END_TYPE

TYPE UDT_DCM :
STRUCT
   Dual_Chanel_Monitor : DCI_MONITOR;
   Status : BOOL;
END_STRUCT
END_TYPE

TYPE UDT_DCS :
STRUCT
   Dual_Chanel_Stop : DCI_STOP;
   Status : BOOL;
END_STRUCT
END_TYPE

TYPE UPS :
STRUCT
   I_Alarm : BOOL;
   I_Battery_Mode : BOOL;
   I_Battery_Charge : BOOL;
   O_Control : BOOL;
END_STRUCT
END_TYPE

TYPE WallClockTimeType :
STRUCT
   Year : DINT;
   Month : DINT;
   Day : DINT;
   Hour : DINT;
   Minute : DINT;
   Second : DINT;
   Microsecond : DINT;
END_STRUCT
END_TYPE

ADD_ON_INSTRUCTION AlarmFallLogUnixon_Dword   (* revision 1.0 *)
VAR_INPUT
   Word_ptr : DINT; {required}
   FallEdge : DINT; {required}
END_VAR
VAR_IN_OUT
   MasterQueue : MasterRTUQueue; {required}
   AssetConfig : AssetSettings; {required}
   FallEvent : SERVER_Interface_RTUData; {required}
END_VAR
VAR
   Bit : DINT; {access None}
END_VAR

ROUTINE Logic   (* ladder *)